(* Logix 5000 project; controller MV vendor 1 type 14 code 217 rev 31.11; software revision 31.00; part 38 of 53 *)
(* tags used below, declared in another part *)
   CWD : CHECKWORD_FLAGS;
   MV_BM01_ZS04 : PlantItem;   // BM01ZS04
   MV_BM01_ZS04_RawInput : ALIAS FOR Remote_IO:8:I.Data.20;   // BM01ZS04
   MV_BM01_ZS05 : PlantItem;   // BM01ZS05
   MV_BM01_ZS05_RawInput : ALIAS FOR Remote_IO:8:I.Data.21;   // BM01ZS05
   MV_FP01_ZS01 : PlantItem;   // FP01ZS01
   MV_FP01_ZS01_RawInput : ALIAS FOR Remote_IO:8:I.Data.16;   // FP01ZS01
   MV_FP01_ZS02 : PlantItem;   // FP01ZS02
   MV_FP01_ZS02_RawInput : ALIAS FOR Remote_IO:8:I.Data.17;   // FP01ZS02
   MV_FP01_ZS03 : PlantItem;   // FP01ZS03
   MV_FP01_ZS03_RawInput : ALIAS FOR Remote_IO:8:I.Data.18;   // FP01ZS03
   MV_FP01_ZS06 : PlantItem;   // FP01ZS06
   MV_FP01_ZS06_RawInput : ALIAS FOR Remote_IO:8:I.Data.19;   // FP01ZS06
   MV_FP01_ZS07 : PlantItem;   // FP01ZS07
   MV_FP01_ZS07_RawInput : ALIAS FOR Remote_IO:8:I.Data.22;   // FP01ZS07
   MV_FP01_ZS08 : PlantItem;   // FP01ZS08
   MV_FP01_ZS08_RawInput : ALIAS FOR Remote_IO:8:I.Data.23;   // FP01ZS08
   MV_MV10_CV1 : PlantItem;   // MV10_CV1
   MV_MV10_CV1_RawOutput : ALIAS FOR Remote_IO:11:O.Data.9;   // MV_MV10_CV1 MV10 coolant SOV
   MV_MV11_CV1 : PlantItem;   // MV11_CV1
   MV_MV11_CV1_RawOutput : ALIAS FOR Remote_IO:11:O.Data.10;   // MV_MV11_CV1 MV11 coolant SOV
   MV_MV12_CV1 : PlantItem;   // MV12_CV1
   MV_MV12_CV1_RawOutput : ALIAS FOR Remote_IO:11:O.Data.11;   // MV_MV12_CV1 MV12 coolant SOV
   MV_MV13_CV1 : PlantItem;   // MV13_CV1
   MV_MV13_CV1_RawOutput : ALIAS FOR Remote_IO:11:O.Data.12;   // MV_MV13_CV1 MV13 coolant SOV
   MV_MV14_CV1 : PlantItem;   // MV14_CV1
   MV_MV14_CV1_RawOutput : ALIAS FOR Remote_IO:11:O.Data.13;   // MV_MV14_CV1 MV14 coolant SOV
   MV_MV15_CV1 : PlantItem;   // MV15_CV1
   MV_MV15_CV1_RawOutput : ALIAS FOR Remote_IO:11:O.Data.14;   // MV_MV15_CV1 MV15 coolant SOV
   MV_MV16_CV1 : PlantItem;   // MV16_CV1
   MV_MV16_CV1_RawOutput : ALIAS FOR Remote_IO:11:O.Data.15;   // MV_MV16_CV1 MV16 coolant SOV
   MV_MV17_CV1 : PlantItem;   // MV17_CV1
   MV_MV17_CV1_RawOutput : ALIAS FOR Remote_IO:12:O.Data.0;   // MV_MV17_CV1 MV17 coolant SOV
   MV_MV18_CV1 : PlantItem;   // MV18_CV1
   MV_MV18_CV1_RawOutput : ALIAS FOR Remote_IO:12:O.Data.1;   // MV_MV18_CV1
   MV_MV19_CV1 : PlantItem;   // MV19_CV1
   MV_MV19_CV1_RawOutput : ALIAS FOR Remote_IO:12:O.Data.2;   // MV_MV19_CV1 MV19 coolant SOV
   MV_MV1_CV1 : PlantItem;   // MV1_CV1
   MV_MV1_CV1_RawOutput : ALIAS FOR Remote_IO:11:O.Data.0;   // MV_MV1_CV1 MV1 coolant SOV
   MV_MV20_CV1 : PlantItem;   // MV20_CV1
   MV_MV20_CV1_RawOutput : ALIAS FOR Remote_IO:12:O.Data.9;   // MV_MV20_CV1 MV23 coolant SOV
   MV_MV21_CV1 : PlantItem;   // MV21_CV1
   MV_MV21_CV1_RawOutput : ALIAS FOR Remote_IO:12:O.Data.10;   // MV_MV21_CV1 MV21coolant SOV
   MV_MV22_CV1 : PlantItem;   // MV22_CV1
   MV_MV22_CV1_RawOutput : ALIAS FOR Remote_IO:12:O.Data.11;   // MV_MV22_CV1 MV22 coolant SOV
   MV_MV23_CV1 : PlantItem;   // MV23_CV1
   MV_MV23_CV1_RawOutput : ALIAS FOR Remote_IO:12:O.Data.12;   // MV_MV23_CV1 MV23 coolant SOV
   MV_MV2_CV1 : PlantItem;   // MV2_CV1
   MV_MV2_CV1_RawOutput : ALIAS FOR Remote_IO:11:O.Data.1;   // MV_MV2_CV1
   MV_MV30_CV1 : PlantItem;   // MV30_CV1
   MV_MV30_CV1_RawOutput : ALIAS FOR Remote_IO:12:O.Data.3;   // MV_MV30_CV1 MV30 coolant SOV
   MV_MV31_CV1 : PlantItem;   // MV31_CV1
   MV_MV31_CV1_RawOutput : ALIAS FOR Remote_IO:12:O.Data.4;   // MV_MV31_CV1 MV31coolant SOV
   MV_MV32_CV1 : PlantItem;   // MV32_CV1
   MV_MV32_CV1_RawOutput : ALIAS FOR Remote_IO:12:O.Data.5;   // MV_MV32_CV1 MV32 coolant SOV
   MV_MV33_CV1 : PlantItem;   // MV33_CV1
   MV_MV33_CV1_RawOutput : ALIAS FOR Remote_IO:12:O.Data.6;   // MV_MV33_CV1 MV33 coolant SOV
   MV_MV34_CV1 : PlantItem;   // MV34_CV1
   MV_MV34_CV1_RawOutput : ALIAS FOR Remote_IO:12:O.Data.7;   // MV_MV34_CV1 MV34 coolant SOV
   MV_MV35_CV1 : PlantItem;   // MV35_CV1
   MV_MV35_CV1_RawOutput : ALIAS FOR Remote_IO:12:O.Data.8;   // MV_MV35_CV1 MV35 coolant SOV
   MV_MV36_AV01 : PlantItem;   // MV36_AV01
   MV_MV36_AV01_RawOutput : ALIAS FOR Remote_IO:16:O.Data.0;   // MV_MV36_AV01
   MV_MV3_CV1 : PlantItem;   // MV3_CV1
   MV_MV3_CV1_RawOutput : ALIAS FOR Remote_IO:11:O.Data.2;   // MV_MV3_CV1 MV3 coolant SOV
   MV_MV4_CV1 : PlantItem;   // MV4_CV1
   MV_MV4_CV1_RawOutput : ALIAS FOR Remote_IO:11:O.Data.3;   // MV_MV4_CV1 MV4 coolant SOV
   MV_MV5_CV1 : PlantItem;   // MV5_CV1
   MV_MV5_CV1_RawOutput : ALIAS FOR Remote_IO:11:O.Data.4;   // MV_MV5_CV1 MV5 coolant SOV
   MV_MV6_CV1 : PlantItem;   // MV6_CV1
   MV_MV6_CV1_RawOutput : ALIAS FOR Remote_IO:11:O.Data.5;   // MV_MV6_CV1 MV6 coolant SOV
   MV_MV7_CV1 : PlantItem;   // MV7_CV1
   MV_MV7_CV1_RawOutput : ALIAS FOR Remote_IO:11:O.Data.6;   // MV_MV7_CV1 MV7 coolant SOV
   MV_MV8_CV1 : PlantItem;   // MV8_CV1
   MV_MV8_CV1_RawOutput : ALIAS FOR Remote_IO:11:O.Data.7;   // MV_MV8_CV1 MV8 coolant SOV
   MV_MV9_CV1 : PlantItem;   // MV9_CV1
   MV_MV9_CV1_RawOutput : ALIAS FOR Remote_IO:11:O.Data.8;   // MV_MV9_CV1 MV9 coolant SOV
   MVCT_Proxies_OK : BOOL;
   MVCT_ProxiesCIP_OK : DINT;
   One_Second_One_Scan : ALIAS FOR One_Second_1_scan;
(* MV_Common, continued *)

ROUTINE MV_Digital_Inputs   (* ladder *)
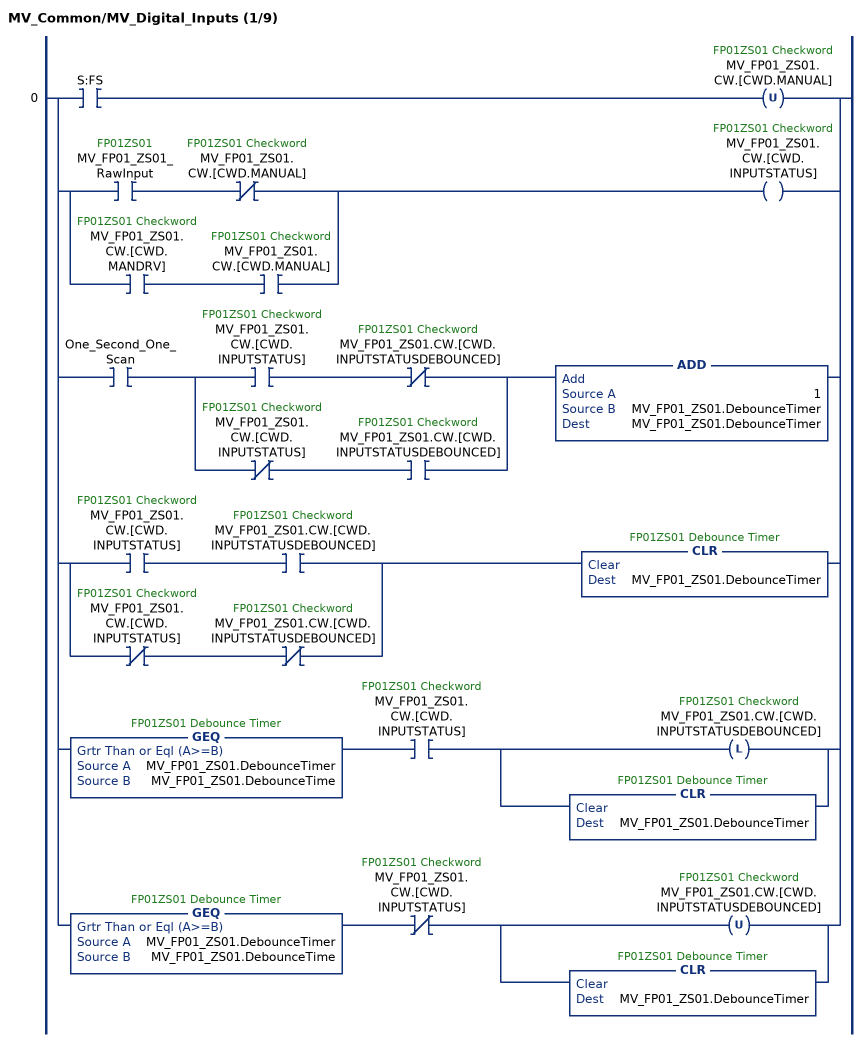
   0: [XIC(S:FS) OTU(MV_FP01_ZS01.CW.[CWD.MANUAL]) ,[XIC(MV_FP01_ZS01_RawInput) XIO(MV_FP01_ZS01.CW.[CWD.MANUAL]) ,XIC(MV_FP01_ZS01.CW.[CWD.MANDRV]) XIC(MV_FP01_ZS01.CW.[CWD.MANUAL]) ] OTE(MV_FP01_ZS01.CW.[CWD.INPUTSTATUS]) ,XIC(One_Second_One_Scan) [XIC(MV_FP01_ZS01.CW.[CWD.INPUTSTATUS]) XIO(MV_FP01_ZS01.CW.[CWD.INPUTSTATUSDEBOUNCED]) ,XIO(MV_FP01_ZS01.CW.[CWD.INPUTSTATUS]) XIC(MV_FP01_ZS01.CW.[CWD.INPUTSTATUSDEBOUNCED]) ] ADD(1,MV_FP01_ZS01.DebounceTimer,MV_FP01_ZS01.DebounceTimer) ,[XIC(MV_FP01_ZS01.CW.[CWD.INPUTSTATUS]) XIC(MV_FP01_ZS01.CW.[CWD.INPUTSTATUSDEBOUNCED]) ,XIO(MV_FP01_ZS01.CW.[CWD.INPUTSTATUS]) XIO(MV_FP01_ZS01.CW.[CWD.INPUTSTATUSDEBOUNCED]) ] CLR(MV_FP01_ZS01.DebounceTimer) ,GEQ(MV_FP01_ZS01.DebounceTimer,MV_FP01_ZS01.DebounceTime) XIC(MV_FP01_ZS01.CW.[CWD.INPUTSTATUS]) [OTL(MV_FP01_ZS01.CW.[CWD.INPUTSTATUSDEBOUNCED]) ,CLR(MV_FP01_ZS01.DebounceTimer) ] ,GEQ(MV_FP01_ZS01.DebounceTimer,MV_FP01_ZS01.DebounceTime) XIO(MV_FP01_ZS01.CW.[CWD.INPUTSTATUS]) [OTU(MV_FP01_ZS01.CW.[CWD.INPUTSTATUSDEBOUNCED]) ,CLR(MV_FP01_ZS01.DebounceTimer) ] ];
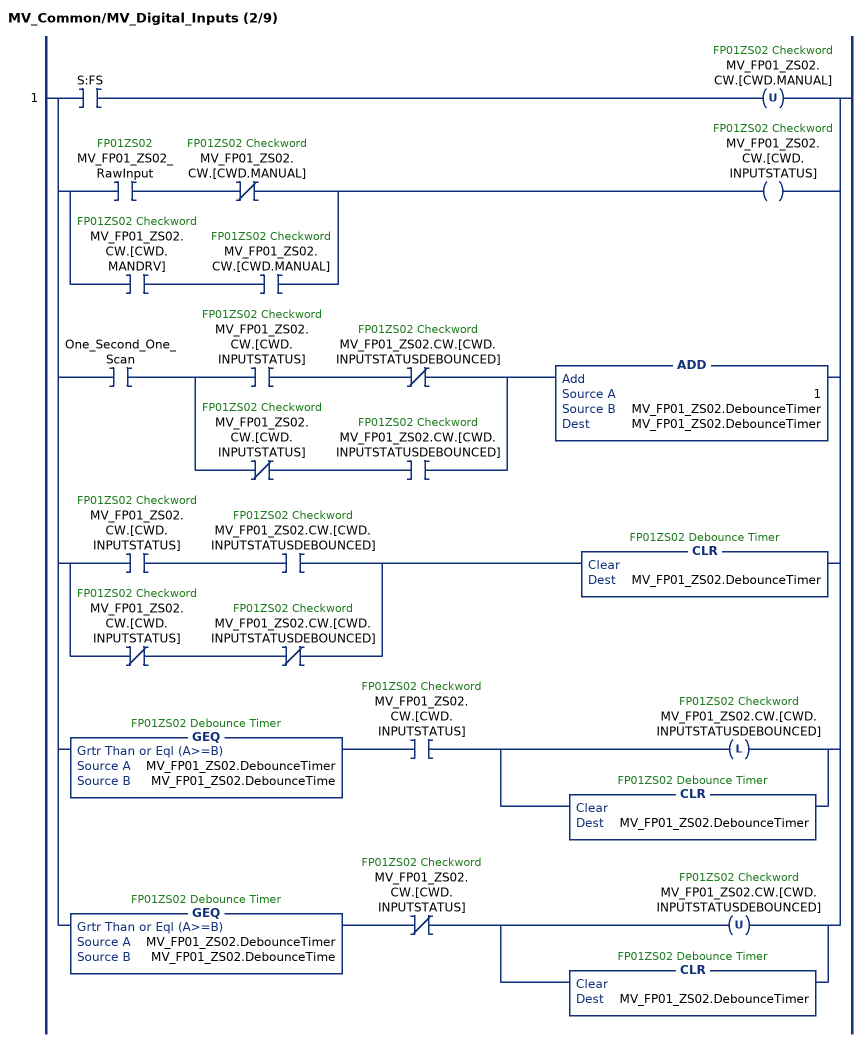
   1: [XIC(S:FS) OTU(MV_FP01_ZS02.CW.[CWD.MANUAL]) ,[XIC(MV_FP01_ZS02_RawInput) XIO(MV_FP01_ZS02.CW.[CWD.MANUAL]) ,XIC(MV_FP01_ZS02.CW.[CWD.MANDRV]) XIC(MV_FP01_ZS02.CW.[CWD.MANUAL]) ] OTE(MV_FP01_ZS02.CW.[CWD.INPUTSTATUS]) ,XIC(One_Second_One_Scan) [XIC(MV_FP01_ZS02.CW.[CWD.INPUTSTATUS]) XIO(MV_FP01_ZS02.CW.[CWD.INPUTSTATUSDEBOUNCED]) ,XIO(MV_FP01_ZS02.CW.[CWD.INPUTSTATUS]) XIC(MV_FP01_ZS02.CW.[CWD.INPUTSTATUSDEBOUNCED]) ] ADD(1,MV_FP01_ZS02.DebounceTimer,MV_FP01_ZS02.DebounceTimer) ,[XIC(MV_FP01_ZS02.CW.[CWD.INPUTSTATUS]) XIC(MV_FP01_ZS02.CW.[CWD.INPUTSTATUSDEBOUNCED]) ,XIO(MV_FP01_ZS02.CW.[CWD.INPUTSTATUS]) XIO(MV_FP01_ZS02.CW.[CWD.INPUTSTATUSDEBOUNCED]) ] CLR(MV_FP01_ZS02.DebounceTimer) ,GEQ(MV_FP01_ZS02.DebounceTimer,MV_FP01_ZS02.DebounceTime) XIC(MV_FP01_ZS02.CW.[CWD.INPUTSTATUS]) [OTL(MV_FP01_ZS02.CW.[CWD.INPUTSTATUSDEBOUNCED]) ,CLR(MV_FP01_ZS02.DebounceTimer) ] ,GEQ(MV_FP01_ZS02.DebounceTimer,MV_FP01_ZS02.DebounceTime) XIO(MV_FP01_ZS02.CW.[CWD.INPUTSTATUS]) [OTU(MV_FP01_ZS02.CW.[CWD.INPUTSTATUSDEBOUNCED]) ,CLR(MV_FP01_ZS02.DebounceTimer) ] ];
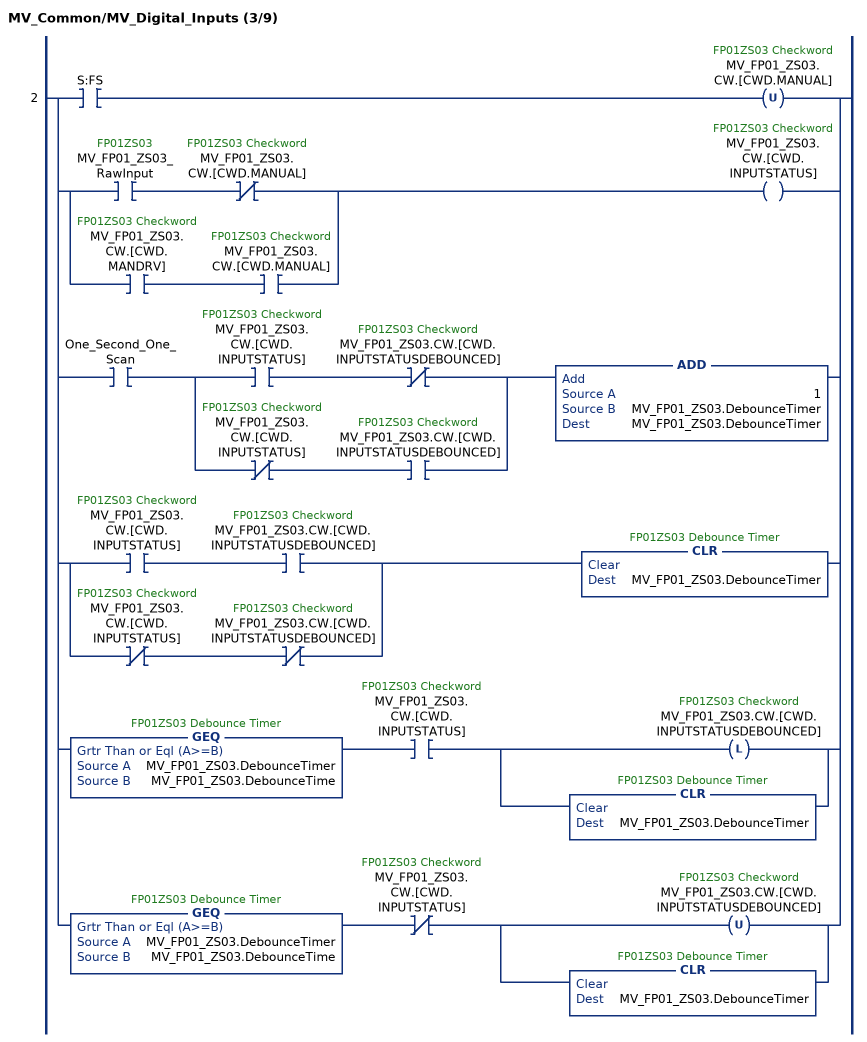
   2: [XIC(S:FS) OTU(MV_FP01_ZS03.CW.[CWD.MANUAL]) ,[XIC(MV_FP01_ZS03_RawInput) XIO(MV_FP01_ZS03.CW.[CWD.MANUAL]) ,XIC(MV_FP01_ZS03.CW.[CWD.MANDRV]) XIC(MV_FP01_ZS03.CW.[CWD.MANUAL]) ] OTE(MV_FP01_ZS03.CW.[CWD.INPUTSTATUS]) ,XIC(One_Second_One_Scan) [XIC(MV_FP01_ZS03.CW.[CWD.INPUTSTATUS]) XIO(MV_FP01_ZS03.CW.[CWD.INPUTSTATUSDEBOUNCED]) ,XIO(MV_FP01_ZS03.CW.[CWD.INPUTSTATUS]) XIC(MV_FP01_ZS03.CW.[CWD.INPUTSTATUSDEBOUNCED]) ] ADD(1,MV_FP01_ZS03.DebounceTimer,MV_FP01_ZS03.DebounceTimer) ,[XIC(MV_FP01_ZS03.CW.[CWD.INPUTSTATUS]) XIC(MV_FP01_ZS03.CW.[CWD.INPUTSTATUSDEBOUNCED]) ,XIO(MV_FP01_ZS03.CW.[CWD.INPUTSTATUS]) XIO(MV_FP01_ZS03.CW.[CWD.INPUTSTATUSDEBOUNCED]) ] CLR(MV_FP01_ZS03.DebounceTimer) ,GEQ(MV_FP01_ZS03.DebounceTimer,MV_FP01_ZS03.DebounceTime) XIC(MV_FP01_ZS03.CW.[CWD.INPUTSTATUS]) [OTL(MV_FP01_ZS03.CW.[CWD.INPUTSTATUSDEBOUNCED]) ,CLR(MV_FP01_ZS03.DebounceTimer) ] ,GEQ(MV_FP01_ZS03.DebounceTimer,MV_FP01_ZS03.DebounceTime) XIO(MV_FP01_ZS03.CW.[CWD.INPUTSTATUS]) [OTU(MV_FP01_ZS03.CW.[CWD.INPUTSTATUSDEBOUNCED]) ,CLR(MV_FP01_ZS03.DebounceTimer) ] ];
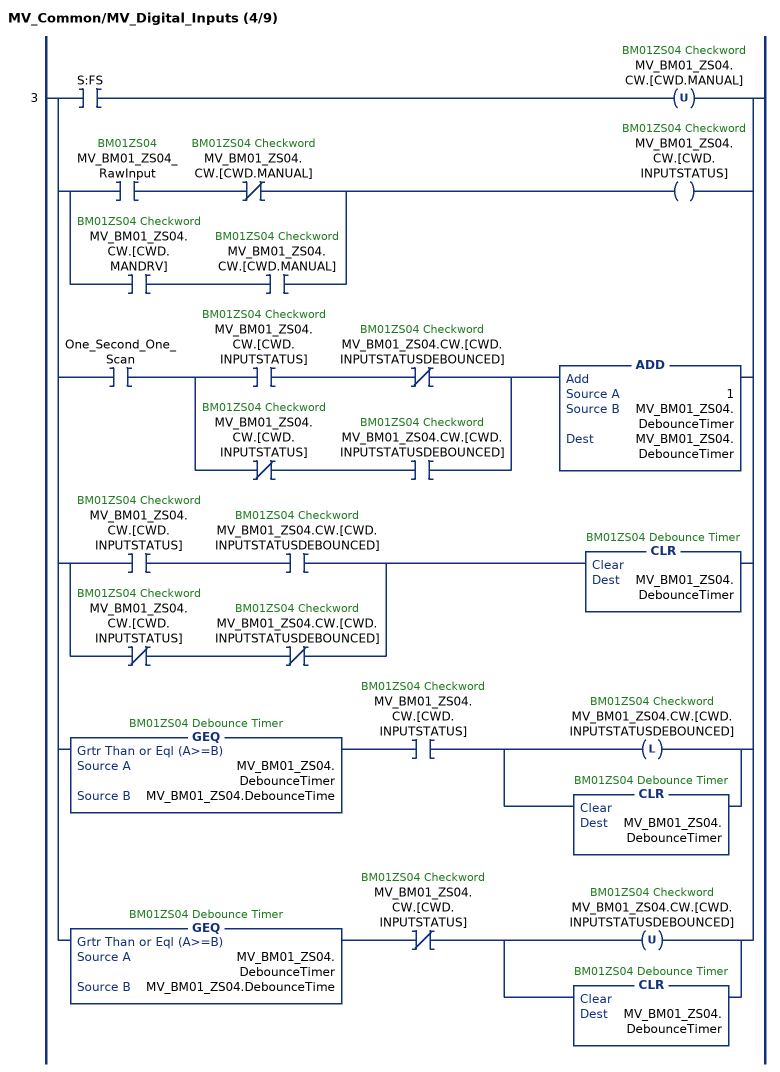
   3: [XIC(S:FS) OTU(MV_BM01_ZS04.CW.[CWD.MANUAL]) ,[XIC(MV_BM01_ZS04_RawInput) XIO(MV_BM01_ZS04.CW.[CWD.MANUAL]) ,XIC(MV_BM01_ZS04.CW.[CWD.MANDRV]) XIC(MV_BM01_ZS04.CW.[CWD.MANUAL]) ] OTE(MV_BM01_ZS04.CW.[CWD.INPUTSTATUS]) ,XIC(One_Second_One_Scan) [XIC(MV_BM01_ZS04.CW.[CWD.INPUTSTATUS]) XIO(MV_BM01_ZS04.CW.[CWD.INPUTSTATUSDEBOUNCED]) ,XIO(MV_BM01_ZS04.CW.[CWD.INPUTSTATUS]) XIC(MV_BM01_ZS04.CW.[CWD.INPUTSTATUSDEBOUNCED]) ] ADD(1,MV_BM01_ZS04.DebounceTimer,MV_BM01_ZS04.DebounceTimer) ,[XIC(MV_BM01_ZS04.CW.[CWD.INPUTSTATUS]) XIC(MV_BM01_ZS04.CW.[CWD.INPUTSTATUSDEBOUNCED]) ,XIO(MV_BM01_ZS04.CW.[CWD.INPUTSTATUS]) XIO(MV_BM01_ZS04.CW.[CWD.INPUTSTATUSDEBOUNCED]) ] CLR(MV_BM01_ZS04.DebounceTimer) ,GEQ(MV_BM01_ZS04.DebounceTimer,MV_BM01_ZS04.DebounceTime) XIC(MV_BM01_ZS04.CW.[CWD.INPUTSTATUS]) [OTL(MV_BM01_ZS04.CW.[CWD.INPUTSTATUSDEBOUNCED]) ,CLR(MV_BM01_ZS04.DebounceTimer) ] ,GEQ(MV_BM01_ZS04.DebounceTimer,MV_BM01_ZS04.DebounceTime) XIO(MV_BM01_ZS04.CW.[CWD.INPUTSTATUS]) [OTU(MV_BM01_ZS04.CW.[CWD.INPUTSTATUSDEBOUNCED]) ,CLR(MV_BM01_ZS04.DebounceTimer) ] ];
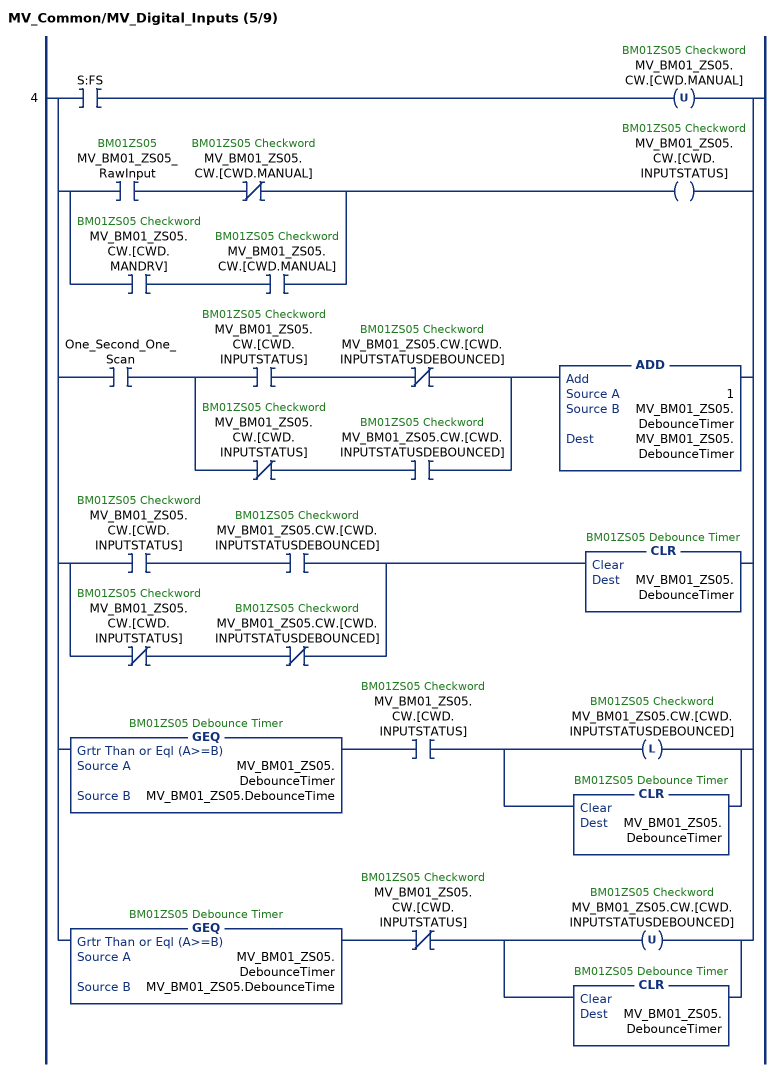
   4: [XIC(S:FS) OTU(MV_BM01_ZS05.CW.[CWD.MANUAL]) ,[XIC(MV_BM01_ZS05_RawInput) XIO(MV_BM01_ZS05.CW.[CWD.MANUAL]) ,XIC(MV_BM01_ZS05.CW.[CWD.MANDRV]) XIC(MV_BM01_ZS05.CW.[CWD.MANUAL]) ] OTE(MV_BM01_ZS05.CW.[CWD.INPUTSTATUS]) ,XIC(One_Second_One_Scan) [XIC(MV_BM01_ZS05.CW.[CWD.INPUTSTATUS]) XIO(MV_BM01_ZS05.CW.[CWD.INPUTSTATUSDEBOUNCED]) ,XIO(MV_BM01_ZS05.CW.[CWD.INPUTSTATUS]) XIC(MV_BM01_ZS05.CW.[CWD.INPUTSTATUSDEBOUNCED]) ] ADD(1,MV_BM01_ZS05.DebounceTimer,MV_BM01_ZS05.DebounceTimer) ,[XIC(MV_BM01_ZS05.CW.[CWD.INPUTSTATUS]) XIC(MV_BM01_ZS05.CW.[CWD.INPUTSTATUSDEBOUNCED]) ,XIO(MV_BM01_ZS05.CW.[CWD.INPUTSTATUS]) XIO(MV_BM01_ZS05.CW.[CWD.INPUTSTATUSDEBOUNCED]) ] CLR(MV_BM01_ZS05.DebounceTimer) ,GEQ(MV_BM01_ZS05.DebounceTimer,MV_BM01_ZS05.DebounceTime) XIC(MV_BM01_ZS05.CW.[CWD.INPUTSTATUS]) [OTL(MV_BM01_ZS05.CW.[CWD.INPUTSTATUSDEBOUNCED]) ,CLR(MV_BM01_ZS05.DebounceTimer) ] ,GEQ(MV_BM01_ZS05.DebounceTimer,MV_BM01_ZS05.DebounceTime) XIO(MV_BM01_ZS05.CW.[CWD.INPUTSTATUS]) [OTU(MV_BM01_ZS05.CW.[CWD.INPUTSTATUSDEBOUNCED]) ,CLR(MV_BM01_ZS05.DebounceTimer) ] ];
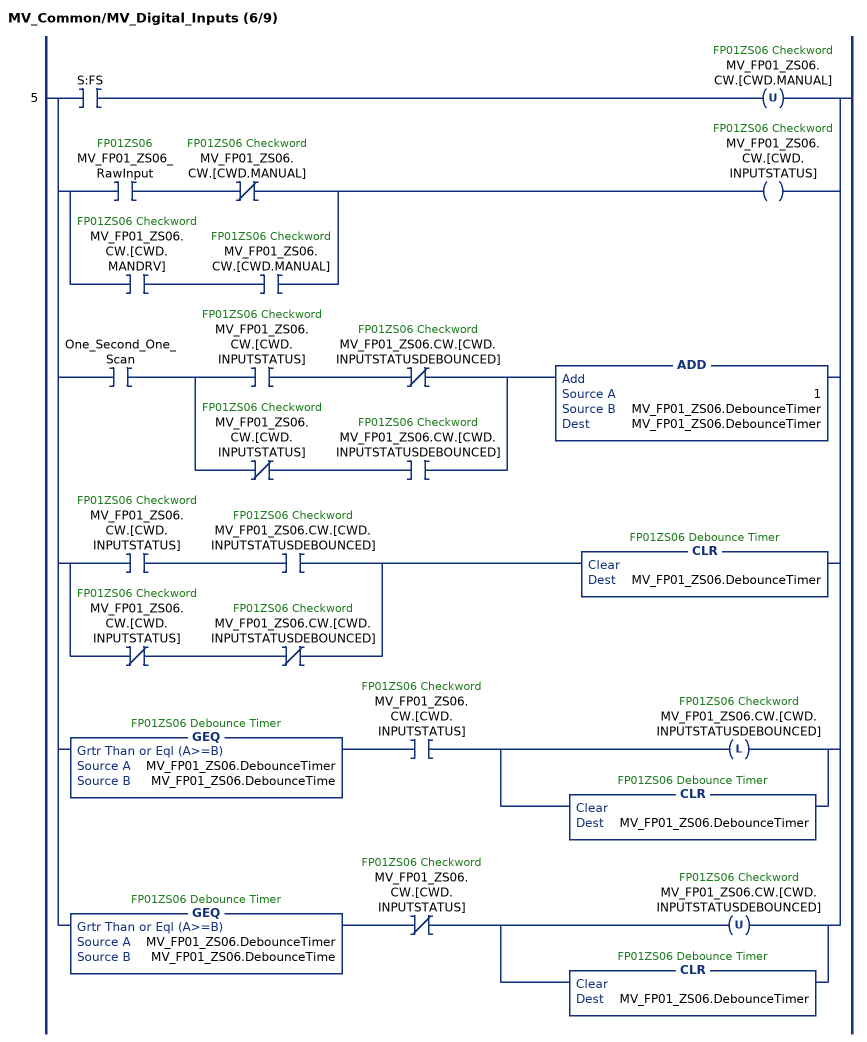
   5: [XIC(S:FS) OTU(MV_FP01_ZS06.CW.[CWD.MANUAL]) ,[XIC(MV_FP01_ZS06_RawInput) XIO(MV_FP01_ZS06.CW.[CWD.MANUAL]) ,XIC(MV_FP01_ZS06.CW.[CWD.MANDRV]) XIC(MV_FP01_ZS06.CW.[CWD.MANUAL]) ] OTE(MV_FP01_ZS06.CW.[CWD.INPUTSTATUS]) ,XIC(One_Second_One_Scan) [XIC(MV_FP01_ZS06.CW.[CWD.INPUTSTATUS]) XIO(MV_FP01_ZS06.CW.[CWD.INPUTSTATUSDEBOUNCED]) ,XIO(MV_FP01_ZS06.CW.[CWD.INPUTSTATUS]) XIC(MV_FP01_ZS06.CW.[CWD.INPUTSTATUSDEBOUNCED]) ] ADD(1,MV_FP01_ZS06.DebounceTimer,MV_FP01_ZS06.DebounceTimer) ,[XIC(MV_FP01_ZS06.CW.[CWD.INPUTSTATUS]) XIC(MV_FP01_ZS06.CW.[CWD.INPUTSTATUSDEBOUNCED]) ,XIO(MV_FP01_ZS06.CW.[CWD.INPUTSTATUS]) XIO(MV_FP01_ZS06.CW.[CWD.INPUTSTATUSDEBOUNCED]) ] CLR(MV_FP01_ZS06.DebounceTimer) ,GEQ(MV_FP01_ZS06.DebounceTimer,MV_FP01_ZS06.DebounceTime) XIC(MV_FP01_ZS06.CW.[CWD.INPUTSTATUS]) [OTL(MV_FP01_ZS06.CW.[CWD.INPUTSTATUSDEBOUNCED]) ,CLR(MV_FP01_ZS06.DebounceTimer) ] ,GEQ(MV_FP01_ZS06.DebounceTimer,MV_FP01_ZS06.DebounceTime) XIO(MV_FP01_ZS06.CW.[CWD.INPUTSTATUS]) [OTU(MV_FP01_ZS06.CW.[CWD.INPUTSTATUSDEBOUNCED]) ,CLR(MV_FP01_ZS06.DebounceTimer) ] ];
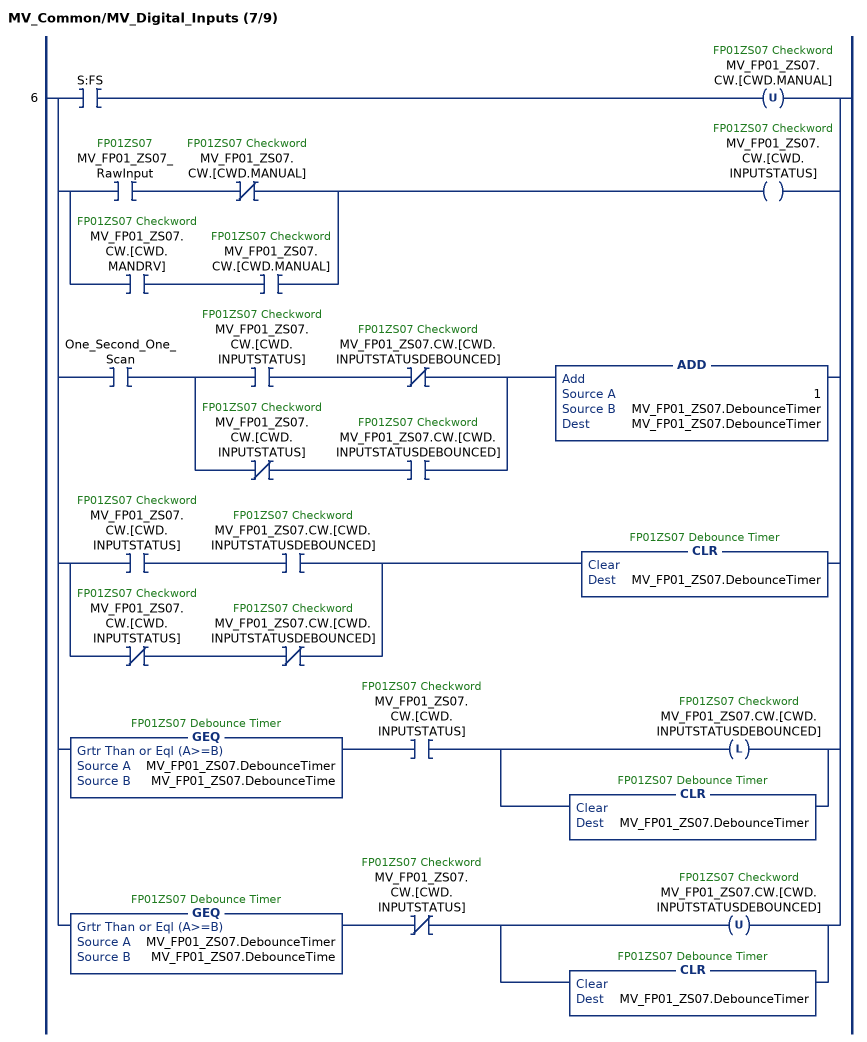
   6: [XIC(S:FS) OTU(MV_FP01_ZS07.CW.[CWD.MANUAL]) ,[XIC(MV_FP01_ZS07_RawInput) XIO(MV_FP01_ZS07.CW.[CWD.MANUAL]) ,XIC(MV_FP01_ZS07.CW.[CWD.MANDRV]) XIC(MV_FP01_ZS07.CW.[CWD.MANUAL]) ] OTE(MV_FP01_ZS07.CW.[CWD.INPUTSTATUS]) ,XIC(One_Second_One_Scan) [XIC(MV_FP01_ZS07.CW.[CWD.INPUTSTATUS]) XIO(MV_FP01_ZS07.CW.[CWD.INPUTSTATUSDEBOUNCED]) ,XIO(MV_FP01_ZS07.CW.[CWD.INPUTSTATUS]) XIC(MV_FP01_ZS07.CW.[CWD.INPUTSTATUSDEBOUNCED]) ] ADD(1,MV_FP01_ZS07.DebounceTimer,MV_FP01_ZS07.DebounceTimer) ,[XIC(MV_FP01_ZS07.CW.[CWD.INPUTSTATUS]) XIC(MV_FP01_ZS07.CW.[CWD.INPUTSTATUSDEBOUNCED]) ,XIO(MV_FP01_ZS07.CW.[CWD.INPUTSTATUS]) XIO(MV_FP01_ZS07.CW.[CWD.INPUTSTATUSDEBOUNCED]) ] CLR(MV_FP01_ZS07.DebounceTimer) ,GEQ(MV_FP01_ZS07.DebounceTimer,MV_FP01_ZS07.DebounceTime) XIC(MV_FP01_ZS07.CW.[CWD.INPUTSTATUS]) [OTL(MV_FP01_ZS07.CW.[CWD.INPUTSTATUSDEBOUNCED]) ,CLR(MV_FP01_ZS07.DebounceTimer) ] ,GEQ(MV_FP01_ZS07.DebounceTimer,MV_FP01_ZS07.DebounceTime) XIO(MV_FP01_ZS07.CW.[CWD.INPUTSTATUS]) [OTU(MV_FP01_ZS07.CW.[CWD.INPUTSTATUSDEBOUNCED]) ,CLR(MV_FP01_ZS07.DebounceTimer) ] ];
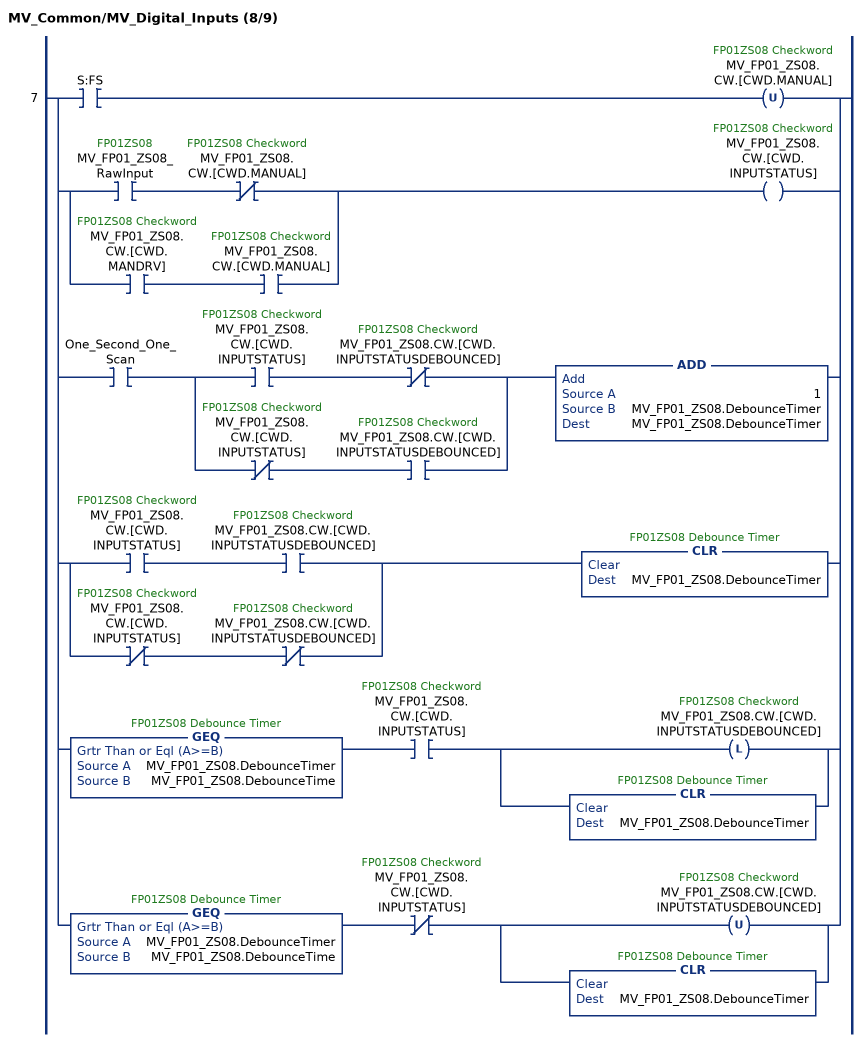
   7: [XIC(S:FS) OTU(MV_FP01_ZS08.CW.[CWD.MANUAL]) ,[XIC(MV_FP01_ZS08_RawInput) XIO(MV_FP01_ZS08.CW.[CWD.MANUAL]) ,XIC(MV_FP01_ZS08.CW.[CWD.MANDRV]) XIC(MV_FP01_ZS08.CW.[CWD.MANUAL]) ] OTE(MV_FP01_ZS08.CW.[CWD.INPUTSTATUS]) ,XIC(One_Second_One_Scan) [XIC(MV_FP01_ZS08.CW.[CWD.INPUTSTATUS]) XIO(MV_FP01_ZS08.CW.[CWD.INPUTSTATUSDEBOUNCED]) ,XIO(MV_FP01_ZS08.CW.[CWD.INPUTSTATUS]) XIC(MV_FP01_ZS08.CW.[CWD.INPUTSTATUSDEBOUNCED]) ] ADD(1,MV_FP01_ZS08.DebounceTimer,MV_FP01_ZS08.DebounceTimer) ,[XIC(MV_FP01_ZS08.CW.[CWD.INPUTSTATUS]) XIC(MV_FP01_ZS08.CW.[CWD.INPUTSTATUSDEBOUNCED]) ,XIO(MV_FP01_ZS08.CW.[CWD.INPUTSTATUS]) XIO(MV_FP01_ZS08.CW.[CWD.INPUTSTATUSDEBOUNCED]) ] CLR(MV_FP01_ZS08.DebounceTimer) ,GEQ(MV_FP01_ZS08.DebounceTimer,MV_FP01_ZS08.DebounceTime) XIC(MV_FP01_ZS08.CW.[CWD.INPUTSTATUS]) [OTL(MV_FP01_ZS08.CW.[CWD.INPUTSTATUSDEBOUNCED]) ,CLR(MV_FP01_ZS08.DebounceTimer) ] ,GEQ(MV_FP01_ZS08.DebounceTimer,MV_FP01_ZS08.DebounceTime) XIO(MV_FP01_ZS08.CW.[CWD.INPUTSTATUS]) [OTU(MV_FP01_ZS08.CW.[CWD.INPUTSTATUSDEBOUNCED]) ,CLR(MV_FP01_ZS08.DebounceTimer) ] ];